		
	10:	// Wait until carrier at stopper
		IF stpStopper.xCarrierAvailable AND NOT xCycleEnd THEN
			uiState := 15;
		END_IF
		
	15:	// Check if RFID tag recognized
		IF stpStopper.dtmRfid.stState.xTagPresent THEN
			uiState := 20;
		ELSE
			uiState := 500;
		END_IF
		
	20:	// Read RFID
		stpStopper.ReadRfid(ADR(stRfidData));
		uiState := 25;
		
	25:	// Wait until read finished
		IF stpStopper.xReady THEN
			uiCarrierId := stRfidData.uiCarrierID;
			uiState := 100;
		END_IF
		
	100:// App. ready and active?
		IF stAppState.xReady AND stAppSettings.xActive THEN
			uiState := 105;
		ELSE
			uiState := 500;
		END_IF
		
	105: // check if carrier already assigned to order
		IF stRfidData.stSapData.udiOp <> udiMyOp AND stRfidData.stSapData.sItem <> 'YE_SMARTMETER' AND xFirstSapModule THEN 			// check if carrier already assigned to order
			SAPInit.Start.Req.sItem := '';
			uiState := 110;
		ELSIF stRfidData.stSapData.udiSfc <> 0 AND stRfidData.stSapData.udiOp = udiMyOp AND stRfidData.stSapData.sItem <> '' THEN		// next operation for this station --> send StartSfc to SAP ME
			udiSfc := stRfidData.stSapData.udiSfc;
			uiState := 200;
		ELSE																															// pass carrier
			uiState := 500;	
		END_IF

///////////////////////////////////
///			 SFC 1010			///
///////////////////////////////////

	110:// Start Sfc (1010)
		xFirstWorkOrder := TRUE;
		SAPInit.Start.Com.iResponse := 0;
		SAPInit.Start.Com.bError	:= FALSE;
		SAPInit.Start.Com.sError	:= '';
        tonHs(IN := FALSE);
        tonOpc(IN := FALSE);
		uiState := 111;
		
		
	111: // Start Sfc Trigger (1010)
		tonOpc(IN := TRUE, PT := T#20MS);
		IF tonOpc.Q THEN
			SAPInit.Start.Com.iTrigger := 1;
			uiState := 115;
		END_IF
		
	115: // Wait Start Sfc (1010) confirmed
		tonHs(IN:= TRUE, PT:= tTimeOutHs);
		IF SAPInit.Start.Com.iTrigger = 0 AND SAPInit.Start.Com.iResponse = 1 THEN
			SAPInit.Start.Com.iResponse := 0;

			IF NOT SAPInit.Start.Com.bError THEN
				uiState := 120;
			ELSE	
				SAPHMI.uiPos  	:= 1; // 1=Start Sfc, 2=Parametric Data, 3=Complete Sfc
				SAPHMI.udiSfc 	:= stRfidData.stSapData.udiSfc;
				SAPHMI.uiOp 	:= stRfidData.stSapData.udiOp;
				SAPHMI.sError	:= SAPInit.Start.Com.sError;
				SAPInit.Start.Com.iTrigger := 0;				
				uiRetryState	:= 110;	
				uiState := 999;
			END_IF
			
		ELSIF tonHs.Q THEN
			SAPHMI.uiPos  	:= 1; // 1=Start Sfc, 2=Parametric Data, 3=Complete Sfc
			SAPHMI.udiSfc 	:= 0;
			SAPHMI.uiOp 	:= stRfidData.stSapData.udiOp;
			SAPHMI.sError	:= 'Handshake timeout';
			SAPInit.Start.Com.iTrigger := 0;
			uiRetryState	:= 110;	
			uiState := 999;
		END_IF
		
	120: // Complete Sfc  (1010)		
		udiSfc := STRING_TO_UDINT(SAPInit.Start.Res.sSfc);
		tonHs(IN:= FALSE);
		IF SAPInit.Start.Res.sItem <> '' AND udiSfc <> 0 THEN
			SAPInit.Comp.Req.sSfc			:= SAPInit.Start.Res.sSfc;
			SAPInit.Comp.Com.iResponse		:= 0;
			SAPInit.Comp.Com.bError			:= FALSE;
			SAPInit.Comp.Com.sError			:= '';
			tonOpc(IN := FALSE);
			uiState := 121;
		ELSE
			uiState := 500;
		END_IF

	121: // Complete Sfc Trigger (1010)
		tonOpc(IN := TRUE, PT := T#20MS);
		IF tonOpc.Q THEN
			SAPInit.Comp.Com.iTrigger := 1;
			uiState := 125;
		END_IF		

	
	125: // Wait Complete Sfc (1010) confirmed
		tonHs(IN := TRUE, PT := tTimeOutHs);
		IF SAPInit.Comp.Com.iTrigger = 0 AND SAPInit.Comp.Com.iResponse = 1 THEN
			SAPInit.Comp.Com.iResponse := 0;
			
			IF NOT SAPInit.Comp.Com.bError THEN
				uiState := 130;
			ELSE	
				SAPHMI.uiPos  	:= 3; // 1=Start Sfc, 2=Parametric Data, 3=Complete Sfc
				SAPHMI.udiSfc 	:= stRfidData.stSapData.udiSfc;
				SAPHMI.uiOp 	:= stRfidData.stSapData.udiOp;
				SAPHMI.sError	:= SAPInit.Comp.Com.sError;
				SAPInit.Comp.Com.iTrigger 		:= 0;
				uiRetryState	:= 120;
				uiState := 999;
			END_IF
			
		ELSIF tonHs.Q THEN
			SAPHMI.uiPos  	:= 3; // 1=Start Sfc, 2=Parametric Data, 3=Complete Sfc
			SAPHMI.udiSfc 	:= 0;
			SAPHMI.uiOp 	:= stRfidData.stSapData.udiOp;
			SAPHMI.sError	:= 'Handshake timeout';
			SAPInit.Comp.Com.iTrigger 		:= 0;
			uiRetryState	:= 120;
			uiState := 999;
		END_IF

	130: // check received operation
		udiOp := STRING_TO_UDINT(SAPInit.Comp.Res.sOp);
		IF udiOp <> 0 THEN
			stRfidData.stSapData.udiSfc		:= udiSfc;
			stRfidData.stSapData.udiOp		:= udiOp;
			stRfidData.stSapData.sItem		:= SAPInit.Start.Res.sItem;
			stRfidData.stSapData.sItemRev	:= SAPInit.Start.Res.sItemRev;
			stRfidData.stSapData.sSfc		:= SAPInit.Start.Res.sSfc;
			uiState := 135;
		ELSE
			uiState := 500;
		END_IF				
		
	135:// Write RFID Data
		stpStopper.WriteRfid(stRfidData);
		uiState := 140;
		
	140: // RFID write OK?
		IF stpStopper.xReady AND NOT stpStopper.dtmRfid.xTimeout AND udiMyOp <> 0 THEN
			uiState := 105;
		ELSIF stpStopper.xReady THEN
			uiState := 500;
		END_IF		


		
///////////////////////////////////
///			 SFC 10xx			///
///////////////////////////////////		

		
	200: // Start Sfc (10xx)		
		xFirstWorkOrder := FALSE;
		SAP.Start.Req.sSfc		:= stRfidData.stSapData.sSfc;
		SAP.Start.Req.sItem		:= stRfidData.stSapData.sItem;
		SAP.Start.Com.iResponse	:= 0;
		SAP.Start.Com.bError	:= FALSE;
		SAP.Start.Com.sError	:= '';
		tonHs(IN := FALSE);
		tonOpc(IN := FALSE);
		uiState	:= 201;
		
		
	201: // Start sfc trigger (10xx)
		tonOpc(In := TRUE, PT := T#20MS);
		IF tonOpc.Q THEN
			SAP.Start.Com.iTrigger := 1;
			tonOpc(IN := FALSE);
			uiState := 205;
		END_IF
		
		
	205: // Wait Start Sfc (10xx) confirmed
		tonHs(IN := TRUE, PT := tTimeOutHs);
		IF SAP.Start.Com.iTrigger = 0 AND SAP.Start.Com.iResponse = 1 THEN
			SAP.Start.Com.iResponse := 0;
			
			IF NOT SAP.Start.Com.bError THEN
				uiState := 220;
			ELSE	
				SAPHMI.uiPos  	:= 1; // 1=Start Sfc, 2=Parametric Data, 3=Complete Sfc
				SAPHMI.udiSfc 	:= stRfidData.stSapData.udiSfc;
				SAPHMI.uiOp 	:= stRfidData.stSapData.udiOp;
				SAPHMI.sError	:= SAP.Start.Com.sError;
				SAP.Start.Com.iTrigger 	:= 0;
				uiRetryState	:= 200;
				uiState := 999;
			END_IF
			
		ELSIF tonHs.Q THEN
			SAPHMI.uiPos  	:= 1; // 1=Start Sfc, 2=Parametric Data, 3=Complete Sfc
			SAPHMI.udiSfc 	:= 0;
			SAPHMI.uiOp 	:= stRfidData.stSapData.udiOp;
			SAPHMI.sError	:= 'Handshake timeout';
			SAP.Start.Com.iTrigger 	:= 0;
			uiRetryState	:= 200;
			uiState := 999;
		END_IF
	
		
	220: // write application parameter
		abySapParameter[0] := SAP.Start.Res.iValue1;
		abySapParameter[1] := SAP.Start.Res.iValue2;	
		abySapParameter[2] := SAP.Start.Res.iValue3;	
		abySapParameter[3] := SAP.Start.Res.iValue4;
		uiState := 300;		
	
				
///////////////////////////////////
///		Start application		///
///////////////////////////////////	

		
	300:// Wait app. free
		IF stAppSettings.xActive AND stAppState.xReady THEN
			uiState := 305;
		END_IF
		
	305:// Send parameters to app 
		stAppControl.auiPar[0] :=	INT_TO_UINT(abySapParameter[0]);
		stAppControl.auiPar[1] :=   INT_TO_UINT(abySapParameter[1]);
		stAppControl.auiPar[2] :=   INT_TO_UINT(abySapParameter[2]);
		stAppControl.auiPar[3] :=   INT_TO_UINT(abySapParameter[3]);
		uiState := 325;
		
	325:// Trigger App. start
		IF stAppSettings.xStopBelt THEN
			convConveyor.Stop();
		END_IF
		stAppControl.xStart := TRUE;
		uiState := 328;
		
	328:// Wait for App. started	
		IF NOT stAppState.xReady THEN
			stAppControl.xStart := FALSE;
			uiState := 330;
		END_IF
		
	330:// Wait for App. finished
		IF stAppState.xReady THEN
			convConveyor.RunToRight(FALSE);
			uiState := 335;
		END_IF
		
	335:// App. fininshed without error?
		IF stAppState.uiReturnCode = 0 THEN
			uiState := 337;
		ELSE
			uiState := 336;
		END_IF
		
	336:// Interactive message
		Visu.stInteractiveError.xError := TRUE;
		Visu.stInteractiveError.sMessageID := UINT_TO_STRING(stAppState.uiReturnCode);
		visu.stInteractiveError.uiAbortState := 337;
		visu.stInteractiveError.uiIgnoreState := 337;
		
		// Retry
		IF visu.stInteractiveError.xBtnRepeat THEN
			visu.stInteractiveError.xBtnRepeat := FALSE;
			visu.stInteractiveError.xError := FALSE;
			uiState := 325;
		END_IF
		
		// Ignore
		IF visu.stInteractiveError.xBtnIgnore THEN
			visu.stInteractiveError.xBtnIgnore := FALSE;
			visu.stInteractiveError.xError := FALSE;
			uiState := visu.stInteractiveError.uiIgnoreState;
		END_IF
		
		// Abort
		IF visu.stInteractiveError.xBtnAbort THEN
			visu.stInteractiveError.xBtnAbort := FALSE;
			visu.stInteractiveError.xError := FALSE;
			uiState := visu.stInteractiveError.uiAbortState;
		END_IF
		
		// Reject order
		IF visu.stInteractiveError.xBtnRejectOrder THEN
			visu.stInteractiveError.xBtnRejectOrder := FALSE;
			visu.stInteractiveError.xError := FALSE;
			uiState := 480;
		END_IF		

///	Paremeters
		
	337: // parametric data
	
		IF xParametricData THEN
			
			IF stAppState.xError THEN
				SAP.Par.Req.iCamResult := 0;
			ELSE
				SAP.Par.Req.iCamResult := 1;
			END_IF
		
		
			SAP.Par.Req.sSfc			:= stRfidData.stSapData.sSfc;
			SAP.Par.Req.sDcGroup		:= SAP.Start.Res.sDcGroup;
			SAP.Par.Req.iValue1			:= SAP.Start.Res.iValue1;
			SAP.Par.Req.sName1			:= SAP.Start.Res.sName1;
			SAP.Par.Req.iValue2			:= SAP.Start.Res.iValue2;
			SAP.Par.Req.sName2			:= SAP.Start.Res.sName2;
			SAP.Par.Req.iValue3			:= SAP.Start.Res.iValue3;
			SAP.Par.Req.sName3			:= SAP.Start.Res.sName3;
			SAP.Par.Req.iValue4			:= SAP.Start.Res.iValue4;
			SAP.Par.Req.sName4			:= SAP.Start.Res.sName4;
			SAP.Par.Com.iResponse		:= 0;
			SAP.Par.Com.bError			:= FALSE;
			SAP.Par.Com.sError			:= '';
        	
			tonHs(In := FALSE);
			tonOpc(In := FALSE);
			uiState := 338;
		ELSE
			uiState := 340;
		END_IF	

	338: // parametric data trigger (10xx)
		tonOpc(In := TRUE, PT := T#20MS);
		IF tonOpc.Q THEN
			SAP.Par.Com.iTrigger := 1;
			tonOpc(IN := FALSE);
			uiState := 339;
		END_IF

	339: // Wait Start Sfc (10xx) confirmed
		tonHs(IN := TRUE, PT := tTimeOutHs);
		IF SAP.Par.Com.iTrigger = 0 AND SAP.Par.Com.iResponse = 1 THEN
			SAP.Par.Com.iResponse := 0;
			
			IF NOT SAP.Par.Com.bError THEN
				uiState := 340;
			ELSE	
				SAPHMI.uiPos  	:= 2; // 1=Start Sfc, 2=Parametric Data, 3=Complete Sfc
				SAPHMI.udiSfc 	:= stRfidData.stSapData.udiSfc;
				SAPHMI.uiOp 	:= stRfidData.stSapData.udiOp;
				SAPHMI.sError	:= SAP.Start.Com.sError;
				SAP.Par.Com.iTrigger 		:= 0;
				uiRetryState	:= 337;
				uiState := 999;
			END_IF
			
		ELSIF tonHs.Q THEN
			SAPHMI.uiPos  	:= 2; // 1=Start Sfc, 2=Parametric Data, 3=Complete Sfc
			SAPHMI.udiSfc 	:= 0;
			SAPHMI.uiOp 	:= stRfidData.stSapData.udiOp;
			SAPHMI.sError	:= 'Handshake timeout';
			SAP.Par.Com.iTrigger 		:= 0;
			uiRetryState	:= 337;
			uiState := 999;
		END_IF		
		
		
		
///	Complete Sfc		
		
	340: // Complete Sfc (10xx)
		SAP.Comp.Req.sSfc		:= stRfidData.stSapData.sSfc;
		SAP.Comp.Com.iResponse	:= 0;
		SAP.Comp.Com.bError		:= FALSE;
		SAP.Comp.Com.sError		:= '';
		
		tonHs(In := FALSE);
		tonOpc(In := FALSE);
		uiState := 341;

	341: // Complete Sfc trigger (10xx)
		tonOpc(In := TRUE, PT := T#20MS);
		IF tonOpc.Q THEN
			SAP.Comp.Com.iTrigger := 1;
			tonOpc(IN := FALSE);
			uiState := 345;
		END_IF

	345: // Wait Complete Sfc (10xx) confirmed
		tonHs(IN := TRUE, PT := tTimeOutHs);
		IF SAP.Comp.Com.iTrigger = 0 AND SAP.Comp.Com.iResponse = 1 THEN
			SAP.Comp.Com.iResponse := 0;
			
			IF NOT SAP.Comp.Com.bError THEN
				uiState := 350;
			ELSE	
				SAPHMI.uiPos  	:= 3; // 1=Start Sfc, 2=Parametric Data, 3=Complete Sfc
				SAPHMI.udiSfc 	:= stRfidData.stSapData.udiSfc;
				SAPHMI.uiOp 	:= stRfidData.stSapData.udiOp;
				SAPHMI.sError	:= SAP.Comp.Com.sError;
				SAP.Comp.Com.iTrigger 	:= 0;
				uiRetryState	:= 340;
				uiState := 999;
			END_IF
			
		ELSIF tonHs.Q THEN
			SAPHMI.uiPos  	:= 3; // 1=Start Sfc, 2=Parametric Data, 3=Complete Sfc
			SAPHMI.udiSfc 	:= 0;
			SAPHMI.uiOp 	:= stRfidData.stSapData.udiOp;
			SAPHMI.sError	:= 'Handshake timeout';
			SAP.Comp.Com.iTrigger 	:= 0;
			uiRetryState	:= 340;
			uiState := 999;
		END_IF
		
	350: //check received operation
		udiOp := STRING_TO_UDINT(SAP.Comp.Res.sOp);
		stRfidData.stSapData.udiOp := udiOp;
		IF udiOp = 0 THEN
			stRfidData.stSapData.udiSfc		:= 0;
			stRfidData.stSapData.sItem		:= '';
			stRfidData.stSapData.sItemRev	:= '';
			stRfidData.stSapData.sSfc		:= '';
		END_IF
		uiState := 400;

		
(*		
	399: // prepare RFID data

		stRfidData.stSapData.udiSfc := 0;
		stRfidData.stSapData.udiOp	:= 0;
		IF stRfidData.stSapData.sItem <> 'YE_SMARTMETER' THEN
			stRfidData.stSapData.sItem := '';
			stRfidData.stSapData.sItemRev := '';
		END_IF
		stRfidData.stSapData.sSfc := '';
		uiState := 400;
*)		
		
		
	400:// Write RFID Data
		stpStopper.WriteRfid(stRfidData);
		uiState := 410;
		
	410:// RFID write OK?
		IF stpStopper.xReady  THEN
			uiState := 500;
		END_IF

		
	500:// Pass carrier
		IF NOT xSemaIn THEN
			xSemaOut := TRUE;
			SAP.Par.Req.sName1		:= '';
			SAP.Par.Req.iValue1		:= 0;
			SAP.Par.Req.sName2		:= '';
			SAP.Par.Req.iValue2		:= 0;
			SAP.Par.Req.sName3		:= '';
			SAP.Par.Req.iValue3		:= 0;
			SAP.Par.Req.sName4		:= '';
			SAP.Par.Req.iValue4		:= 0;
			SAP.Par.Req.sDcGroup	:= '';
			stpStopper.Release();
			uiState := 505;
		END_IF
		
	505:// Wait for release
		IF stpStopper.xReady THEN
			uiState := 10;
		END_IF
		
	999:// Interactive message
		Visu.stInteractiveError.xError := TRUE;
		visu.stInteractiveError.uiAbortState := 350;
		
		// Retry
		IF visu.stInteractiveError.xBtnRepeat THEN
			visu.stInteractiveError.xBtnRepeat := FALSE;
			visu.stInteractiveError.xError := FALSE;
			uiState := uiRetryState;
		END_IF
	
		// Abort
		IF visu.stInteractiveError.xBtnAbort THEN
			visu.stInteractiveError.xBtnAbort := FALSE;
			visu.stInteractiveError.xError := FALSE;
			uiState := visu.stInteractiveError.uiAbortState;
		END_IF
		
		
	
END_CASE
END_METHOD

END_FUNCTION_BLOCK

// Programs/SwitchWithoutMes
FUNCTION_BLOCK SwitchWithoutMes
VAR_INPUT
	byMode				: BYTE;
	uiResourceId		: UINT := 0;
	usiCanNodeId		: USINT := 33;
	usiCanNetworkId		: USINT := 0;
	usiCanChannel		: USINT := 1;
	udiMyOp				: UDINT;

	xRfid_SiemensByteOrder: BOOL;
	xCarrierAvSensor: BOOL;
	xCarrierIdBit0: BOOL;
	xCarrierIdBit1: BOOL;
	xCarrierIdBit2: BOOL;
	xStopperReleased: BOOL;
	xSwitchInByPassDir: BOOL;
	xSwitchInStraightDir:BOOL;
	xTraficSensorStraight: BOOL;
	xTrafficSensorByPass: BOOL;
END_VAR
VAR_OUTPUT
	xInitPos			: BOOL;
	xLeft				: BOOL;
	xRight				: BOOL;
	xSlow				: BOOL;
	xStop				: BOOL;
	stAppControl		: st_AppControl;
	stAppSettings		: st_AppSettings;

	xReleaseStopper		: BOOL;
	xSwitchToByPass		: BOOL;
	xSwitchToStraight	: BOOL;
END_VAR
VAR_IN_OUT
	astTransitionTable	: ARRAY [0..10] OF st_TransitionData;
END_VAR
VAR
	uiState				: UINT := 0;
	convConveyor		: dc_ecp.Conveyor2Dir;
	stpStopper			: dc_ecp.CPF_StopperDtm425;
	stRfidData			: dc_ecp.st_CPF_RfidData;
	xFirstWorkOrder		: BOOL := FALSE;
	udiONo				: UDINT;
	uiOPos				: UINT;
	uiOpNo				: UINT;
	uiCarrierId			: UINT;
	ftAuto				: F_TRIG;
	ftManual			: F_TRIG;
	uiActualTransitionRow: UINT;
	uiNextState: UINT;
	uiI: UINT;
	xValidOperation: BOOL;
	uiCarrierInitNum	: UINT;
	uiCondIn		: UINT;
	uiCondOut		: UINT;
	xSwitch: BOOL;
END_VAR


////////////////////////////////////////////
// Execute moduls
////////////////////////////////////////////

_ModuleCalls();

		
////////////////////////////////////////////
// Init RFID
////////////////////////////////////////////
IF NOT stpStopper.xConnected AND stpStopper.xReady THEN	
	stpStopper.Connect(usiCanNodeId:= usiCanNodeId, usiCanNetworkId:= usiCanNetworkId, usiCanChannel:= usiCanChannel);
END_IF


////////////////////////////////////////////
// MES Mode
////////////////////////////////////////////

// Execute MES mode
IF xAuto AND byMode = 1 THEN
	_MesMode();
END_IF



////////////////////////////////////////////
// Exit from auto or manual mode
////////////////////////////////////////////

ftAuto(CLK := xAuto);
ftManual(CLK := xManual);

IF ftAuto.Q OR ftManual.Q THEN
	convConveyor.Stop();
	stpStopper.cpfssStopper.MoveUp();
	uiState := 0;
END_IF


xInitPos := (uiState <= 10);

////////////////////////////////////////////
// Default Mode
////////////////////////////////////////////

// Execute Default Mode
IF xAuto AND byMode = 0 THEN
	_DefaultMode();
END_IF

////////////////////////////////////////////
// SAP Mode
////////////////////////////////////////////

// Execute SAP Mode
IF xAuto AND byMode = 2 THEN
	_SapMode();
END_IF

METHOD PRIVATE _SapMode : BOOL
VAR_INPUT
END_VAR
CASE uiState OF
	0:	// Idle
		convConveyor.Stop();
		IF xAuto THEN
			uiState := 1;
		END_IF
		
	1:	// Init
		convConveyor.RunToRight(FALSE);
		uiState := 2;
		
	2:	// Wait for RFID
		IF stpStopper.xReady AND stpStopper.xConnected THEN
			uiState := 10;
		END_IF
		
	10:	// Wait until carrier at stopper
		IF stpStopper.xCarrierAvailable AND NOT xCycleEnd THEN
			xSwitch := FALSE;
			uiState := 15;
		END_IF
		
	15:	// Check if RFID tag recognized
		IF stpStopper.dtmRfid.stState.xTagPresent THEN
			uiState := 20;
		ELSE
			uiState := 500;
		END_IF
		
	20:	// Read RFID
		stpStopper.ReadRfid(ADR(stRfidData));
		uiState := 25;
		
	25:	// Wait until read finished
		IF stpStopper.xReady THEN
			uiState := 300;
		END_IF
		
	300:// Change the switch variable
		IF stRfidData.stSapData.udiOp = udiMyOp THEN
			xSwitch := TRUE;			
		END_IF
		
		uiState := 490;
		
	490:// Change the switch
		IF xSwitch AND NOT xTrafficSensorByPass THEN
			xSwitch := TRUE;
			xSwitchToByPass := TRUE;
			xSwitchToStraight := FALSE;	
			uiState := 495;	
		ELSIF NOT xTraficSensorStraight THEN
			xSwitch := FALSE;
			xSwitchToByPass := FALSE;
			xSwitchToStraight := TRUE;	
			uiState := 495;	
		END_IF

	495:// Wait for Switch
		IF (NOT xSwitch AND xSwitchInStraightDir) OR (XSwitch AND xSwitchInByPassDir) THEN
			uiState := 500;
		END_IF
		
	500:// Pass carrier
		IF (xSwitch AND NOT xTrafficSensorByPass) OR (NOT xSwitch AND NOT xTraficSensorStraight) THEN
			stpStopper.Release();
			uiState := 505;
		END_IF
		
	505:// Wait for release
		IF stpStopper.xReady THEN
			uiState := 510;
		END_IF
		
	510://Wait for trafic
		IF (xSwitch AND xTrafficSensorByPass) OR (NOT xSwitch AND xTraficSensorStraight) THEN
			uiState := 10;
		END_IF
	
END_CASE
END_METHOD

METHOD PRIVATE _MesMode : BOOL
VAR_INPUT
END_VAR
VAR
END_VAR
CASE uiState OF
	0:	// Idle
		convConveyor.Stop();
		IF xAuto THEN
			uiState := 1;
		END_IF
		
	1:	// Wait for RFID
		IF stpStopper.xReady AND stpStopper.xConnected THEN
			convConveyor.RunToRight(FALSE);
			uiState := 10;
		END_IF		

		
	10:	// Wait until carrier at stopper
		IF stpStopper.xCarrierAvailable AND NOT xCycleEnd THEN
			xSwitch := FALSE;
			uiState := 15;
		END_IF
		
	15:	// Check if RFID tag recognized
		IF stpStopper.dtmRfid.stState.xTagPresent THEN
			uiState := 20;
		ELSE
			uiState := 500;
		END_IF
		
	20:	// Read RFID
		stpStopper.ReadRfid(ADR(stRfidData));
		uiState := 25;
		
	25:	// Wait until read finished
		IF stpStopper.xReady THEN
			uiState := 300;
		END_IF
		
	300:// Change the switch variable
		IF stRfidData.stMesData.uiResourceId = uiResourceId THEN
			xSwitch := TRUE;			
		END_IF
		
		uiState := 490;
		
	490:// Change the switch
		IF xSwitch AND NOT xTrafficSensorByPass THEN
			xSwitch := TRUE;
			xSwitchToByPass := TRUE;
			xSwitchToStraight := FALSE;	
			uiState := 495;	
		ELSIF NOT xTraficSensorStraight THEN
			xSwitch := FALSE;
			xSwitchToByPass := FALSE;
			xSwitchToStraight := TRUE;	
			uiState := 495;	
		END_IF

	495:// Wait for Switch
		IF (NOT xSwitch AND xSwitchInStraightDir) OR (XSwitch AND xSwitchInByPassDir) THEN
			uiState := 500;
		END_IF
		
	500:// Pass carrier
		IF (xSwitch AND NOT xTrafficSensorByPass) OR (NOT xSwitch AND NOT xTraficSensorStraight) THEN
			stpStopper.Release();
			uiState := 505;
		END_IF
		
	505:// Wait for release
		IF stpStopper.xReady THEN
			uiState := 510;
		END_IF
		
	510://Wait for trafic
		IF (xSwitch AND xTrafficSensorByPass) OR (NOT xSwitch AND xTraficSensorStraight) THEN
			uiState := 10;
		END_IF
	
END_CASE
END_METHOD

METHOD PRIVATE _DefaultMode : BOOL
VAR_INPUT
END_VAR
VAR
END_VAR
CASE uiState OF
	0:	// Idle
		convConveyor.Stop();
		IF xAuto THEN
			uiState := 1;
		END_IF
		
	1:	// Init
		convConveyor.RunToRight(FALSE);
		uiState := 2;
		
	2:	// Wait for RFID
		IF stpStopper.xReady AND stpStopper.xConnected THEN
			uiState := 10;
		END_IF
		
	10:	// Wait until carrier at stopper
		IF stpStopper.xCarrierAvailable AND NOT xCycleEnd THEN
			xSwitch := FALSE;
			uiState := 15;
		END_IF
		
	15:	// Check if RFID tag recognized
		IF stpStopper.dtmRfid.stState.xTagPresent THEN
			uiState := 20;
		ELSE
			uiState := 500;
		END_IF
		
	20:	// Read RFID
		stpStopper.ReadRfid(ADR(stRfidData));
		uiState := 25;
		
	25:	// Wait until read finished
		IF stpStopper.xReady THEN
			uiState := 50;
		END_IF
		
	50:	// check carrier init condition
		IF stAppSettings.xCarrierInit THEN
			uiCondIn := 0;
			uiCondOut := astTransitionTable[0].uiCondOut;
			uiState := 55;
		ELSE
			// TODO: "dbAppPar".Init.iCntAct := 0; ???
			uiState := 65;
		END_IF
		
	55:	// check if Application is enabled in init step
		uiCarrierInitNum := uiCarrierInitNum + 1;
		IF uiCarrierInitNum >= stAppSettings.uiCarrierInitNum THEN
			uiCarrierInitNum := 0;
			stAppSettings.xCarrierInit := FALSE;
		END_IF	
	
		IF astTransitionTable[0].xAppEn THEN
			uiActualTransitionRow := 0;
			uiState := 300;
		ELSE
			
			SysMemSet(pDest := ADR(stRfidData.stMesData), udiValue := 0, udiCount := SIZEOF(stRfidData.stMesData));
			stRfidData.uiCode := astTransitionTable[0].uiCondOut;
			// TODO: "dbAppPar".Init.iCntAct := "dbAppPar".Init.iCntAct + 1;
			uiState := 400;
			
		END_IF

	65:	// Check application start condition
        uiNextState := 490;
		
		// Search for a raw with the input condition
		uiCondIn := stRfidData.uiCode;
		uiCondOut := 0;
        FOR uiI := 1 TO 10 DO
            IF (uiCondIn = astTransitionTable[uiI].uiCondIn) AND (stRfidData.uiCode <> 0) THEN
				//Entry condition o.k.
                IF astTransitionTable[uiI].xAppEn THEN
                    // application for this condition activated
					uiActualTransitionRow := uiI;
					uiCondOut := astTransitionTable[uiI].uiCondOut;
                    uiNextState := 300;
                    EXIT;
                ELSE
                    // no application start, only write output code to RFID
                    stRfidData.uiCode := astTransitionTable[uiI].uiCondOut;
                    uiNextState := 400;
                    EXIT;
                END_IF
            END_IF
        END_FOR
		
        uiState := uiNextState;
		
	300:// Change the switch variable
		IF astTransitionTable[uiActualTransitionRow].uiPar1 <> 0 THEN
			xSwitch := TRUE;			
		END_IF
		
		stRfidData.uiCode := astTransitionTable[uiActualTransitionRow].uiCondOut;	
		uiState := 400;
				
	400:// Write RFID Data
		stpStopper.WriteRfid(stRfidData);
		uiState := 410;
		
	410:// Wait RFID write finished
		IF stpStopper.xReady THEN
			uiState := 490;
		END_IF
		
	490:// Change the switch
		IF xSwitch AND NOT xTrafficSensorByPass THEN
			xSwitch := TRUE;
			xSwitchToByPass := TRUE;
			xSwitchToStraight := FALSE;	
			uiState := 495;	
		ELSIF NOT xTraficSensorStraight THEN
			xSwitch := FALSE;
			xSwitchToByPass := FALSE;
			xSwitchToStraight := TRUE;
			uiState := 495;		
		END_IF
		
	495:// Wait for Switch
		IF (NOT xSwitch AND xSwitchInStraightDir) OR (XSwitch AND xSwitchInByPassDir) THEN
			uiState := 500;
		END_IF
		
	500:// Pass carrier
		IF (xSwitch AND NOT xTrafficSensorByPass) OR (NOT xSwitch AND NOT xTraficSensorStraight) THEN
			stpStopper.Release();
			uiState := 505;
		END_IF
		
	505:// Wait for release
		IF stpStopper.xReady THEN
			uiState := 510;
		END_IF
		
	510://Wait for trafic
		IF (xSwitchInByPassDir AND xTrafficSensorByPass) OR (xSwitchInStraightDir AND xTraficSensorStraight) THEN
			uiState := 10;
		END_IF
	
	
END_CASE
END_METHOD

METHOD PRIVATE _ModuleCalls : BOOL
VAR_INPUT
END_VAR
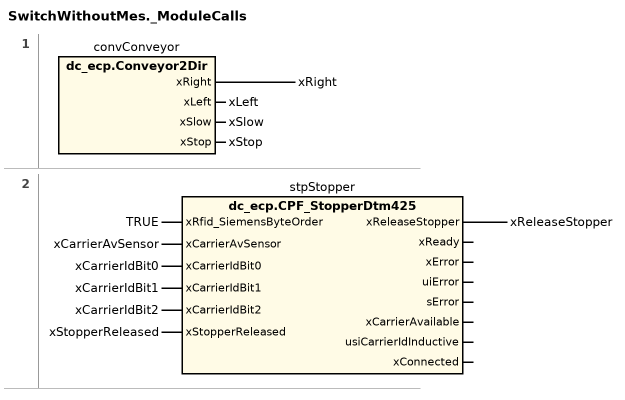
// NETWORK 1
convConveyor(xLeft => xLeft, xSlow => xSlow, xStop => xStop); // dc_ecp.Conveyor2Dir
xRight := convConveyor.xRight;

// NETWORK 2
stpStopper(
    xRfid_SiemensByteOrder := TRUE,
    xCarrierAvSensor := xCarrierAvSensor,
    xCarrierIdBit0 := xCarrierIdBit0,
    xCarrierIdBit1 := xCarrierIdBit1,
    xCarrierIdBit2 := xCarrierIdBit2,
    xStopperReleased := xStopperReleased); // dc_ecp.CPF_StopperDtm425
xReleaseStopper := stpStopper.xReleaseStopper;
END_METHOD

END_FUNCTION_BLOCK

// Programs/Tools/ErrorCpyHMI
PROGRAM ErrorCpyHMI
VAR
	///Rising edges for write
	artWritingEdge: ARRAY[0..191] OF R_TRIG;
	///Rising edges for delete
	aftDeletingEdge: ARRAY[0..191] OF F_TRIG;
	///Variable for the FOR loop
	uiI: UINT;
	///Pointer to the errors
	pbError: POINTER TO BYTE;
END_VAR

//------------------------------------------------------------------------
// Handle the date for the HMI
//------------------------------------------------------------------------


FOR uiI := 0 TO 191 DO			//There are 64 errors in 3 level (3*64 = 192, /0 --> 191/)

//------------------------------------------------------------------------
// Checking the errors
//------------------------------------------------------------------------	
	pbError := ADR(stError) + (uiI/8);
	artWritingEdge[uiI](CLK := (pbError^ AND SHL(1,uiI MOD 8)) > 0 );	
	aftDeletingEdge[uiI](CLK := (pbError^ AND SHL(1,uiI MOD 8)) > 0 );	
	
//Write into the error table
	IF artWritingEdge[uiI].Q THEN
			Visu.fbErrorFifo.sErrorID := CONCAT('L', CONCAT(UINT_TO_STRING((uiI) / 64), CONCAT('.', UINT_TO_STRING((uiI) MOD 64))));  
			Visu.fbErrorFifo(xWrite := FALSE);
			Visu.fbErrorFifo(xWrite := TRUE);
	END_IF
	
//Delete from the error table
	IF aftDeletingEdge[uiI].Q THEN
			Visu.fbErrorFifo.sErrorID := CONCAT('L', CONCAT(UINT_TO_STRING((uiI) / 64), CONCAT('.', UINT_TO_STRING((uiI) MOD 64))));  
			Visu.fbErrorFifo(xDelete := FALSE);
			Visu.fbErrorFifo(xDelete := TRUE);
	END_IF
	
END_FOR

END_PROGRAM

// Programs/Tools/ErrorCpyWinCC
PROGRAM ErrorCpyWinCC
VAR
	/// number of bytes to copy
	udiCount: UDINT;
	/// Timer to extend the global error flag
	TOF_SF: TOF;
END_VAR

//------------------------------------------------------------------------
// ErrorCpy 
//	- Calculates error WORDs from BITs
//------------------------------------------------------------------------

stError.xSF0 := (stError.uL0.lwError <> 0);
stError.xSF1 := (stError.uL1.lwError <> 0);
stError.xSF2 := (stError.uL2.lwError <> 0);

//----------------------------------------------------------------------------------------------
// summary error flag for LEVEL 0 OR LEVEL 1 errors
//----------------------------------------------------------------------------------------------
stError.xSF := stError.xSF0 OR stError.xSF1;

//----------------------------------------------------------------------------------------------
// extend xSF with 100ms
//----------------------------------------------------------------------------------------------
TOF_SF(IN := stError.xSF, PT:= T#100MS); 
stError.xSF_ext := TOF_SF.Q;

END_PROGRAM

// Programs/SwitchWithMes
FUNCTION_BLOCK SwitchWithMes
VAR_INPUT
	byMode				: BYTE;
	usiCanNodeId		: USINT := 33;
	usiCanNetworkId		: USINT := 0;
	usiCanChannel		: USINT := 1;
	sMesIp				: STRING := '172.20.0.90';
	uiMesQueryPort		: UINT := 2000;
	uiMesStatePort		: UINT := 2001;
	uiResourceId		: UINT := 0;
	stAppState			: st_AppState;
	stAppInfo			: st_AppInfo;
	udiBranchOp				: UDINT;

	xRfid_SiemensByteOrder: BOOL;
	xCarrierAvSensor: BOOL;
	xCarrierIdBit0: BOOL;
	xCarrierIdBit1: BOOL;
	xCarrierIdBit2: BOOL;
	xStopperReleased: BOOL;
	xSwitchInByPassDir: BOOL;
	xSwitchInStraightDir:BOOL;
	xTraficSensorStraight: BOOL;
	xTrafficSensorByPass: BOOL;
	xSemaIn			: BOOL;
END_VAR
VAR_OUTPUT
	xInitPos			: BOOL;
	xLeft				: BOOL;
	xRight				: BOOL;
	xSlow				: BOOL;
	xStop				: BOOL;
	stAppControl		: st_AppControl;
	stAppSettings		: st_AppSettings;

	xReleaseStopper		: BOOL;
	xSwitchToByPass		: BOOL;
	xSwitchToStraight	: BOOL;
	xSemaOut			: BOOL;
END_VAR
VAR_IN_OUT
	astTransitionTable	: ARRAY [0..10] OF st_TransitionData;
END_VAR
VAR
	uiState				: UINT := 0;
	convConveyor		: dc_ecp.Conveyor2Dir;
	stpStopper			: dc_ecp.CPF_StopperDtm425;
	mesMES				: dc_ecp.MES4;
	stRfidData			: dc_ecp.st_CPF_RfidData;
	stRcvHeader			: dc_ecp.st_MES4_QueryHeader;
	auiRcvPar			: ARRAY [0..3] OF UINT;
	auiSndPar			: ARRAY [0..3] OF UINT;
	xFirstWorkOrder		: BOOL := FALSE;
	udiONo				: UDINT;
	uiOPos				: UINT;
	uiOpNo				: UINT;
	uiCarrierId			: UINT;
	ftAuto				: F_TRIG;
	ftManual			: F_TRIG;
	uiActualTransitionRow: UINT;
	uiNextState: UINT;
	uiI: UINT;
	xValidOperation: BOOL;
	uiCarrierInitNum	: UINT;
	uiCondIn		: UINT;
	uiCondOut		: UINT;
	xSwitch: BOOL;
	stShuntId	: st_GetShuntId;
	uiShuntId	: UINT;
END_VAR

xSemaOut := xSemaIn;
////////////////////////////////////////////
// Execute moduls
////////////////////////////////////////////

_ModuleCalls();

		
////////////////////////////////////////////
// Init RFID
////////////////////////////////////////////
IF NOT stpStopper.xConnected AND stpStopper.xReady THEN	
	stpStopper.Connect(usiCanNodeId:= usiCanNodeId, usiCanNetworkId:= usiCanNetworkId, usiCanChannel:= usiCanChannel);
END_IF


////////////////////////////////////////////
// MES Mode
////////////////////////////////////////////

// Execute MES mode
IF xAuto AND byMode = 1 THEN
	_MesMode();
END_IF

// Connect to MES
IF (NOT mesMES.xConnected AND mesMEs.xReady) OR mesMES.xError THEN
	mesMES.Connect(sIP := sMesIp, uiQueryPort := uiMesQueryPort, uiStatePort := uiMesStatePort, uiResourceId := uiResourceId);
END_IF


////////////////////////////////////////////
// Exit from auto or manual mode
////////////////////////////////////////////

ftAuto(CLK := xAuto);
ftManual(CLK := xManual);

IF ftAuto.Q OR ftManual.Q THEN
	convConveyor.Stop();
	stpStopper.cpfssStopper.MoveUp();
	uiState := 0;
END_IF

stAppControl.xReset := xReset;

mesMES.stResourceState.xAuto := xAuto;
mesMES.stResourceState.xManual := xManual;
mesMES.stResourceState.xReset := xReset;
mesMES.stResourceState.xMES := xMES;
mesMES.stResourceState.xErrL0 := stError.xSF0;
mesMES.stResourceState.xErrL1 := stError.xSF1;
mesMES.stResourceState.xErrL2 := stError.xSF2;
mesMES.stResourceState.xBusy := NOT stAppState.xReady;

xInitPos := (uiState <= 10) AND stAppState.xInitPos;


////////////////////////////////////////////
// Default Mode
////////////////////////////////////////////

// Execute Default Mode
IF xAuto AND byMode = 0 THEN
	_DefaultMode();
END_IF

////////////////////////////////////////////
// SAP Mode
////////////////////////////////////////////

// Execute SAP Mode
IF xAuto AND byMode = 2 THEN
	_SapMode();
END_IF

METHOD PRIVATE _DefaultMode : BOOL
VAR_INPUT
END_VAR
VAR
END_VAR
CASE uiState OF
	0:	// Idle
		convConveyor.Stop();
		IF xAuto THEN
			uiState := 1;
		END_IF
		
	1:	// Init
		convConveyor.RunToRight(FALSE);
		uiState := 2;
		
	2:	// Wait for RFID
		IF stpStopper.xReady AND stpStopper.xConnected THEN
			uiState := 10;
		END_IF
		
	10:	// Wait until carrier at stopper
		IF stpStopper.xCarrierAvailable AND NOT xCycleEnd THEN
			xSwitch := FALSE;
			uiState := 15;
		END_IF
		
	15:	// Check if RFID tag recognized
		IF stpStopper.dtmRfid.stState.xTagPresent THEN
			uiState := 20;
		ELSE
			xSwitch := FALSE;
			uiState := 490;
		END_IF
		
	20:	// Read RFID
		stpStopper.ReadRfid(ADR(stRfidData));
		uiState := 25;
		
	25:	// Wait until read finished
		IF stpStopper.xReady THEN
			uiState := 50;
		END_IF
		
	50:	// check carrier init condition
		IF stAppSettings.xCarrierInit THEN
			uiCondIn := 0;
			uiCondOut := astTransitionTable[0].uiCondOut;
			uiState := 55;
		ELSE
			// TODO: "dbAppPar".Init.iCntAct := 0; ???
			uiState := 65;
		END_IF
		
	55:	// check if Application is enabled in init step
		uiCarrierInitNum := uiCarrierInitNum + 1;
		IF uiCarrierInitNum >= stAppSettings.uiCarrierInitNum THEN
			uiCarrierInitNum := 0;
			stAppSettings.xCarrierInit := FALSE;
		END_IF	
	
		IF astTransitionTable[0].xAppEn THEN
			uiActualTransitionRow := 0;
			uiState := 300;
		ELSE
			
			SysMemSet(pDest := ADR(stRfidData.stMesData), udiValue := 0, udiCount := SIZEOF(stRfidData.stMesData));
			stRfidData.uiCode := astTransitionTable[0].uiCondOut;
			// TODO: "dbAppPar".Init.iCntAct := "dbAppPar".Init.iCntAct + 1;
			uiState := 400;
			
		END_IF

	65:	// Check application start condition
        uiNextState := 490;
		
		// Search for a raw with the input condition
		uiCondIn := stRfidData.uiCode;
		uiCondOut := 0;
        FOR uiI := 1 TO 10 DO
            IF (uiCondIn = astTransitionTable[uiI].uiCondIn) AND (stRfidData.uiCode <> 0) THEN
				//Entry condition o.k.
                IF astTransitionTable[uiI].xAppEn THEN
                    // application for this condition activated
					uiActualTransitionRow := uiI;
					uiCondOut := astTransitionTable[uiI].uiCondOut;
                    uiNextState := 300;
                    EXIT;
                ELSE
                    // no application start, only write output code to RFID
                    stRfidData.uiCode := astTransitionTable[uiI].uiCondOut;
                    uiNextState := 400;
                    EXIT;
                END_IF
            END_IF
        END_FOR
		
        uiState := uiNextState;
		
	300:// Change the switch variable
		IF astTransitionTable[uiActualTransitionRow].uiPar1 <> 0 THEN
			xSwitch := TRUE;			
		END_IF
		
		stRfidData.uiCode := astTransitionTable[uiActualTransitionRow].uiCondOut;	
		uiState := 400;
				
	400:// Write RFID Data
		stpStopper.WriteRfid(stRfidData);
		uiState := 410;
		
	410:// Wait RFID write finished
		IF stpStopper.xReady THEN
			uiState := 490;
		END_IF
		
	490:// Change the switch
		IF xSwitch AND NOT xTrafficSensorByPass  THEN
			xSwitchToByPass := TRUE;
			xSwitchToStraight := FALSE;	
			uiState := 495;	
		ELSIF NOT xTraficSensorStraight AND NOT xSemaIn THEN
			xSwitchToByPass := FALSE;
			xSwitchToStraight := TRUE;
			xSemaOut		:= TRUE;
			uiState := 495;		
		END_IF
		
	495:// Wait for Switch
		IF (NOT xSwitch AND xSwitchInStraightDir) OR (XSwitch AND xSwitchInByPassDir) THEN
			uiState := 500;
		END_IF
		
	500:// Pass carrier
		IF (xSwitch AND NOT xTrafficSensorByPass) OR (NOT xSwitch AND NOT xTraficSensorStraight) THEN
			
			stpStopper.Release();
			uiState := 505;
		END_IF
		
	505:// Wait for release
		IF stpStopper.xReady THEN
			uiState := 510;
		END_IF
		
	510://Wait for trafic
		IF (xSwitchInByPassDir AND xTrafficSensorByPass) OR (xSwitchInStraightDir AND xTraficSensorStraight) THEN
			uiState := 10;
		END_IF
	
	
END_CASE
END_METHOD

METHOD PRIVATE _ModuleCalls : BOOL
VAR_INPUT
END_VAR
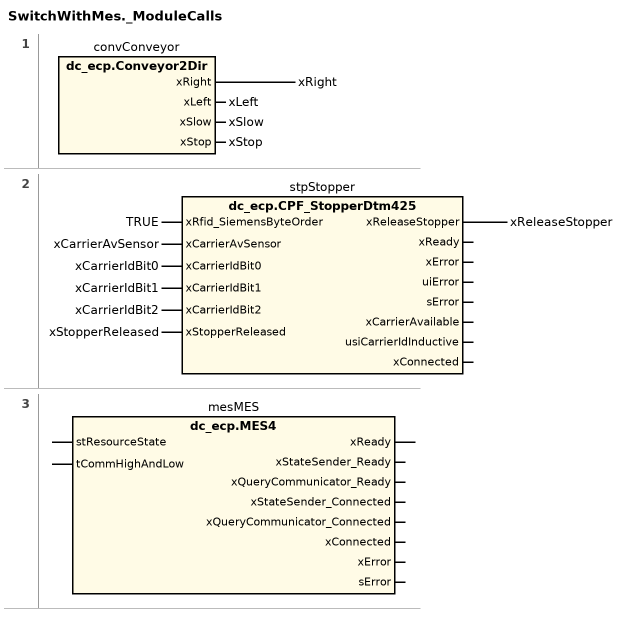
// NETWORK 1
convConveyor(xLeft => xLeft, xSlow => xSlow, xStop => xStop); // dc_ecp.Conveyor2Dir
xRight := convConveyor.xRight;

// NETWORK 2
stpStopper(
    xRfid_SiemensByteOrder := TRUE,
    xCarrierAvSensor := xCarrierAvSensor,
    xCarrierIdBit0 := xCarrierIdBit0,
    xCarrierIdBit1 := xCarrierIdBit1,
    xCarrierIdBit2 := xCarrierIdBit2,
    xStopperReleased := xStopperReleased); // dc_ecp.CPF_StopperDtm425
xReleaseStopper := stpStopper.xReleaseStopper;

// NETWORK 3
mesMES(); // dc_ecp.MES4
END_METHOD

METHOD PRIVATE _SapMode : BOOL
VAR_INPUT
END_VAR
VAR
END_VAR
CASE uiState OF
	0:	// Idle
		convConveyor.Stop();
		IF xAuto THEN
			uiState := 1;
		END_IF
		
	1:	// Init
		convConveyor.RunToRight(FALSE);
		uiState := 2;
		
	2:	// Wait for RFID
		IF stpStopper.xReady AND stpStopper.xConnected THEN
			uiState := 10;
		END_IF
		
	10:	// Wait until carrier at stopper
		IF stpStopper.xCarrierAvailable AND NOT xCycleEnd THEN
			xSwitch := FALSE;
			uiState := 15;
		END_IF
		
	15:	// Check if RFID tag recognized
		IF stpStopper.dtmRfid.stState.xTagPresent THEN
			uiState := 20;
		ELSE
			xSwitch := FALSE;
			uiState := 490;
		END_IF
		
	20:	// Read RFID
		stpStopper.ReadRfid(ADR(stRfidData));
		uiState := 25;
		
	25:	// Wait until read finished
		IF stpStopper.xReady THEN
			uiState := 300;
		END_IF
		
	300:// Change the switch variable
		IF stRfidData.stSapData.udiOp = udiBranchOp THEN
			xSwitch := TRUE;			
		END_IF
		
		uiState := 490;
		
	490:// Change the switch
		IF xSwitch AND NOT xTrafficSensorByPass THEN
			xSwitch := TRUE;
			xSwitchToByPass := TRUE;
			xSwitchToStraight := FALSE;	
			uiState := 495;	
		ELSIF NOT xTraficSensorStraight THEN
			xSwitch := FALSE;
			xSwitchToByPass := FALSE;
			xSwitchToStraight := TRUE;	
			uiState := 495;	
		END_IF

	495:// Wait for Switch
		IF (NOT xSwitch AND xSwitchInStraightDir) OR (XSwitch AND xSwitchInByPassDir) THEN
			uiState := 500;
		END_IF
		
	500:// Pass carrier
		IF (xSwitch AND NOT xTrafficSensorByPass) OR (NOT xSwitch AND NOT xTraficSensorStraight) THEN
			stpStopper.Release();
			uiState := 505;
		END_IF
		
	505:// Wait for release
		IF stpStopper.xReady THEN
			uiState := 510;
		END_IF
		
	510://Wait for trafic
		IF (xSwitch AND xTrafficSensorByPass) OR (NOT xSwitch AND xTraficSensorStraight) THEN
			uiState := 10;
		END_IF
	
END_CASE
END_METHOD

METHOD PRIVATE _MesMode : BOOL
VAR_INPUT
END_VAR
VAR
END_VAR
CASE uiState OF
	0:	// Idle
		convConveyor.Stop();
		IF xAuto THEN
			uiState := 1;
		END_IF
		
	1: // Init
		IF mesMES.xConnected THEN
			convConveyor.RunToRight(FALSE);
			uiState := 2;
		END_IF	
		
		
	2:	// Wait for RFID
		IF stpStopper.xReady AND stpStopper.xConnected THEN
			uiState := 10;
		END_IF
	
		
	10:	// Wait until carrier at stopper
		IF stpStopper.xCarrierAvailable AND NOT xCycleEnd  THEN
			uiState := 15;
		END_IF
		
	15:	// Check if RFID tag recognized
		IF stpStopper.dtmRfid.stState.xTagPresent THEN
			uiState := 20;
		ELSE
			xSwitch := FALSE;
			uiState := 490;
		END_IF
		
	20:	// Read RFID
		stpStopper.ReadRfid(ADR(stRfidData));
		uiState := 25;
		
	25:	// Wait until read finished
		IF stpStopper.xReady THEN
			uiState := 26;
		END_IF
		
	26: //pass empty carriers
		IF stRfidData.stMesData.udiONo = 0 THEN
			xSwitch := FALSE; //empty carriers go straight.
			uiState := 490;
		ELSE
			uiState := 300;				
		END_IF
		
		
	300://  Get this order
		stShuntId.uiSourceId:=uiResourceId;
		stShuntId.uiSourcePosition:=2;
		stShuntId.uiTargetId:=stRfidData.stMesData.uiResourceId;
		stShuntId.uiTargetPosition:=1;
	
		mesMES.GetShuntForTarget(
				pRcvHeader:= ADR(stRcvHeader), 
				pRcvPar:= ADR(uiShuntId), 
				szRcvPar:= SIZEOF(uiShuntId), 
				pSndPar:= ADR(stShuntId), 
				szSndPar:= SIZEOF(stShuntId));
		uiState := 305;
		
	305:// Wait for MES request
		IF stRcvHeader.xDone THEN
			uiState := 310;
		ELSIF xCycleEnd THEN
			uiState := 500;	
		END_IF
	
	310: // Set path
		IF uiShuntId = 2 THEN
			xSwitch		:= TRUE;
		ELSE
			xSwitch		:= FALSE;
		END_IF
		uiState := 490;
		
	490:// Change the switch
		IF xSwitch AND NOT xTrafficSensorByPass  THEN
			xSwitchToByPass := TRUE;
			xSwitchToStraight := FALSE;	
			uiState := 495;	
		ELSIF NOT xTraficSensorStraight AND NOT xSemaIn THEN
			xSwitchToByPass := FALSE;
			xSwitchToStraight := TRUE;
			xSemaOut := TRUE;	
			uiState := 495;	
		END_IF

	495:// Wait for Switch
		IF (NOT xSwitch AND xSwitchInStraightDir) OR (XSwitch AND xSwitchInByPassDir) THEN
			uiState := 500;
		END_IF
		
	500:// Pass carrier
		IF (xSwitch AND NOT xTrafficSensorByPass) OR (NOT xSwitch AND NOT xTraficSensorStraight) THEN
			stpStopper.Release();
			uiState := 505;
		END_IF
		
	505:// Wait for release
		IF stpStopper.xReady THEN
			uiState := 510;
		END_IF
		
	510://Wait for trafic
		IF (xSwitch AND xTrafficSensorByPass) OR (NOT xSwitch AND xTraficSensorStraight) THEN
			uiState := 10;
		END_IF
	
END_CASE
END_METHOD

END_FUNCTION_BLOCK
